// Mitsubishi GX Works2 project: KotelnyaPLC   PLC: FX3U/FX3UC (continued)
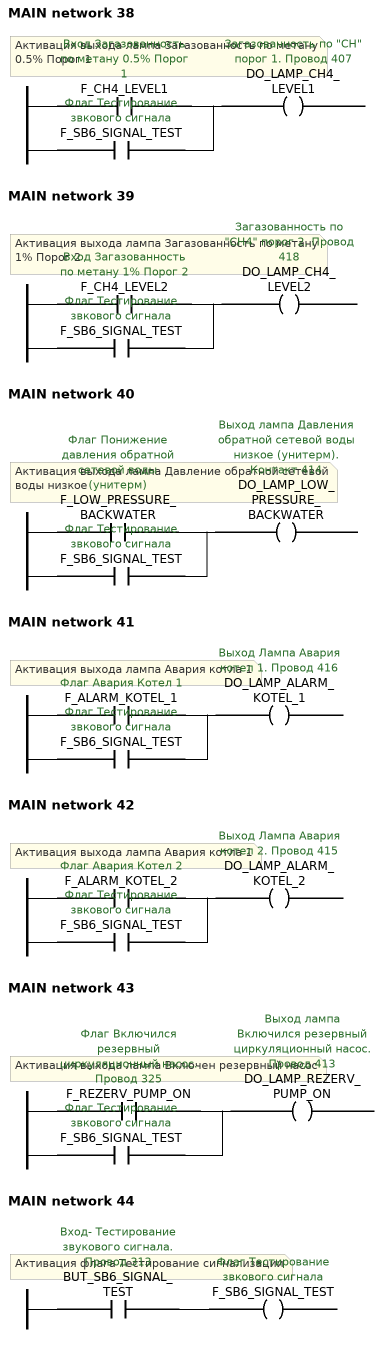
(* [picture p5: structured ladder/FBD of MAIN, networks 38 to 44] *)
(* network 38 *)
(* Активация выхода лампа Загазованность по метану 0.5% Порог 1 *)
DO_LAMP_CH4_LEVEL1 := F_CH4_LEVEL1 OR F_SB6_SIGNAL_TEST;
(* network 39 *)
(* Активация выхода лампа Загазованность по метану 1% Порог 2 *)
DO_LAMP_CH4_LEVEL2 := F_CH4_LEVEL2 OR F_SB6_SIGNAL_TEST;
(* network 40 *)
(* Активация выхода лампа Давление обратной сетевой воды низкое *)
DO_LAMP_LOW_PRESSURE_BACKWATER := F_LOW_PRESSURE_BACKWATER OR F_SB6_SIGNAL_TEST;
(* network 41 *)
(* Активация выхода лампа Авария котла 1 *)
DO_LAMP_ALARM_KOTEL_1 := F_ALARM_KOTEL_1 OR F_SB6_SIGNAL_TEST;
(* network 42 *)
(* Активация выхода лампа Авария котла 1 *)
DO_LAMP_ALARM_KOTEL_2 := F_ALARM_KOTEL_2 OR F_SB6_SIGNAL_TEST;
(* network 43 *)
(* Активация выхода лампа Включен резервный насос *)
DO_LAMP_REZERV_PUMP_ON := F_REZERV_PUMP_ON OR F_SB6_SIGNAL_TEST;
(* network 44 *)
(* Активация флага Тестирование сигнализации *)
F_SB6_SIGNAL_TEST := BUT_SB6_SIGNAL_TEST;
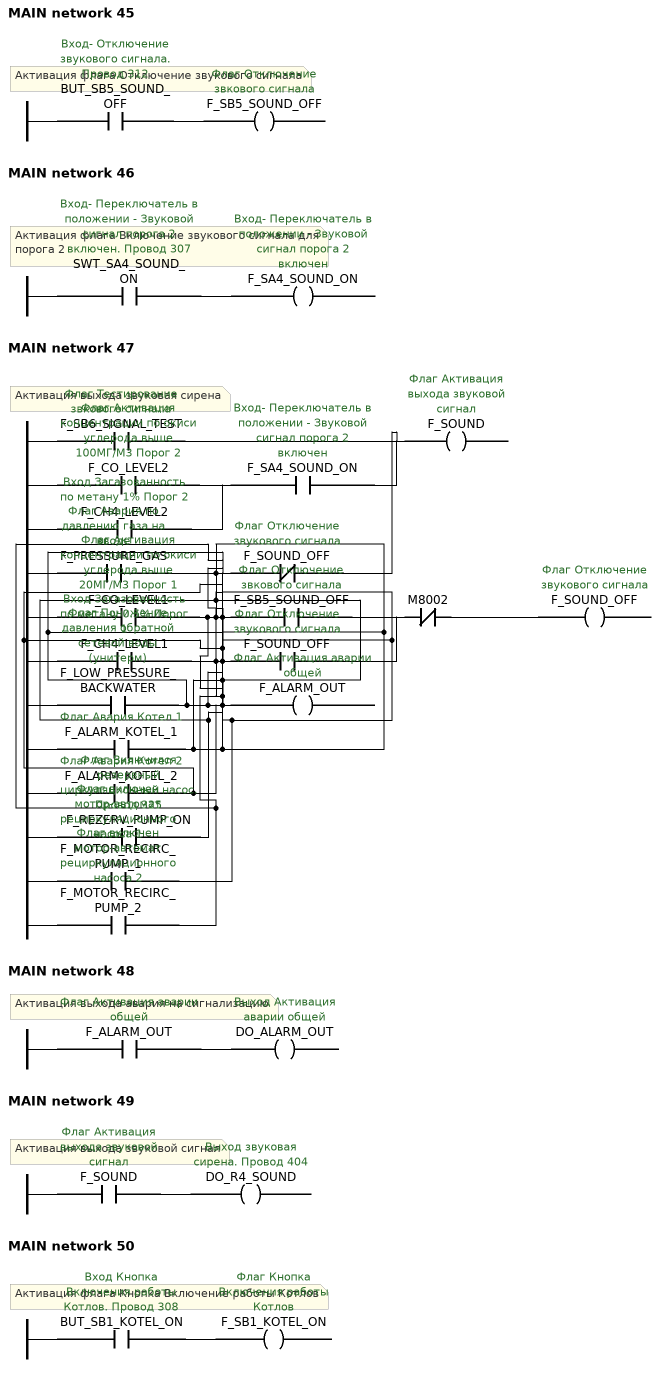
(* network 45 *)
(* Активация флага Отключение звукового сигнала *)
F_SB5_SOUND_OFF := BUT_SB5_SOUND_OFF;
(* network 46 *)
(* Активация флага Включение звукового сигнала для порога 2 *)
F_SA4_SOUND_ON := SWT_SA4_SOUND_ON;
(* network 47 *)
(* Активация выхода звуковая сирена *)
_p1 := F_PRESSURE_GAS OR F_CO_LEVEL1 OR F_CH4_LEVEL1 OR F_LOW_PRESSURE_BACKWATER OR F_ALARM_KOTEL_1 OR F_ALARM_KOTEL_2 OR F_REZERV_PUMP_ON OR F_MOTOR_RECIRC_PUMP_1 OR F_MOTOR_RECIRC_PUMP_2;
F_SOUND := F_SB6_SIGNAL_TEST OR ((F_CO_LEVEL2 OR F_CH4_LEVEL2) AND F_SA4_SOUND_ON) OR (_p1 AND NOT F_SOUND_OFF);
F_SOUND_OFF := ((_p1 AND F_SB5_SOUND_OFF) OR (_p1 AND F_SOUND_OFF)) AND NOT M8002;
F_ALARM_OUT := _p1;
(* network 48 *)
(* Активация выхода авария на сигнализацию *)
DO_ALARM_OUT := F_ALARM_OUT;
(* network 49 *)
(* Активация выхода звуковой сигнал *)
DO_R4_SOUND := F_SOUND;
(* network 50 *)
(* Активация флага Кнопка Включение работы Котлов *)
F_SB1_KOTEL_ON := BUT_SB1_KOTEL_ON;
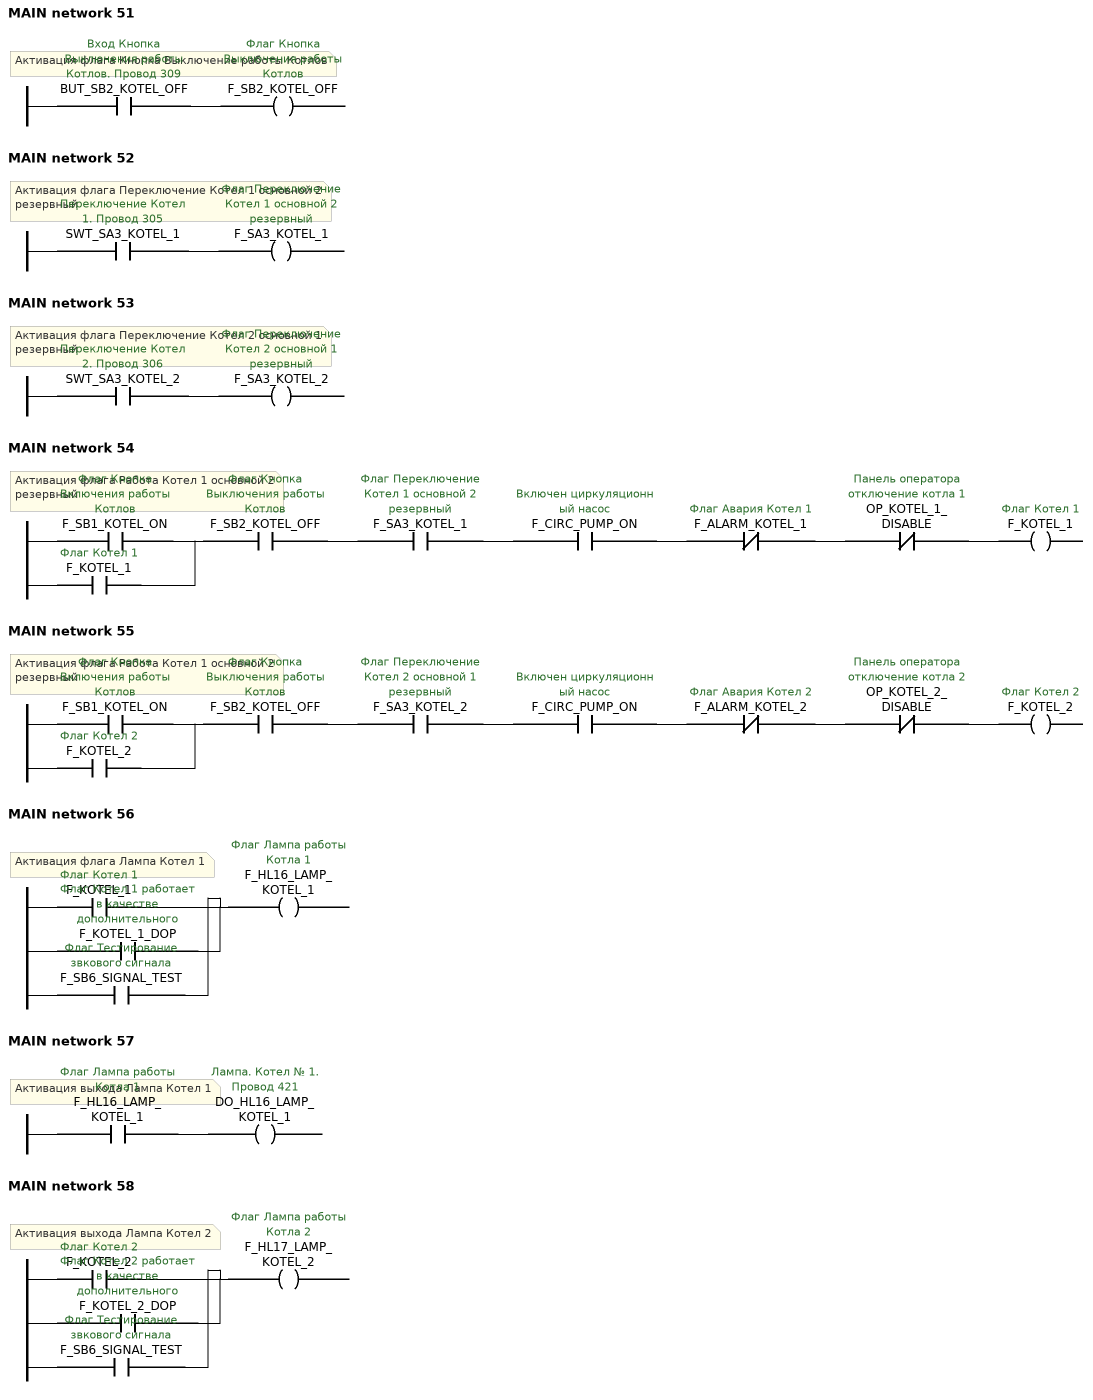
(* network 51 *)
(* Активация флага Кнопка Выключение работы Котлов *)
F_SB2_KOTEL_OFF := BUT_SB2_KOTEL_OFF;
(* network 52 *)
(* Активация флага Переключение Котел 1 основной 2 резервный *)
F_SA3_KOTEL_1 := SWT_SA3_KOTEL_1;
(* network 53 *)
(* Активация флага Переключение Котел 2 основной 1 резервный *)
F_SA3_KOTEL_2 := SWT_SA3_KOTEL_2;
(* network 54 *)
(* Активация флага Работа Котел 1 основной 2 резервный *)
F_KOTEL_1 := (((((F_SB1_KOTEL_ON OR F_KOTEL_1) AND F_SB2_KOTEL_OFF) AND F_SA3_KOTEL_1) AND F_CIRC_PUMP_ON) AND NOT F_ALARM_KOTEL_1) AND NOT OP_KOTEL_1_DISABLE;
(* network 55 *)
(* Активация флага Работа Котел 1 основной 2 резервный *)
F_KOTEL_2 := (((((F_SB1_KOTEL_ON OR F_KOTEL_2) AND F_SB2_KOTEL_OFF) AND F_SA3_KOTEL_2) AND F_CIRC_PUMP_ON) AND NOT F_ALARM_KOTEL_2) AND NOT OP_KOTEL_2_DISABLE;
(* network 56 *)
(* Активация флага Лампа Котел 1 *)
F_HL16_LAMP_KOTEL_1 := F_KOTEL_1 OR F_KOTEL_1_DOP OR F_SB6_SIGNAL_TEST;
(* network 57 *)
(* Активация выхода Лампа Котел 1 *)
DO_HL16_LAMP_KOTEL_1 := F_HL16_LAMP_KOTEL_1;
(* network 58 *)
(* Активация выхода Лампа Котел 2 *)
F_HL17_LAMP_KOTEL_2 := F_KOTEL_2 OR F_KOTEL_2_DOP OR F_SB6_SIGNAL_TEST;
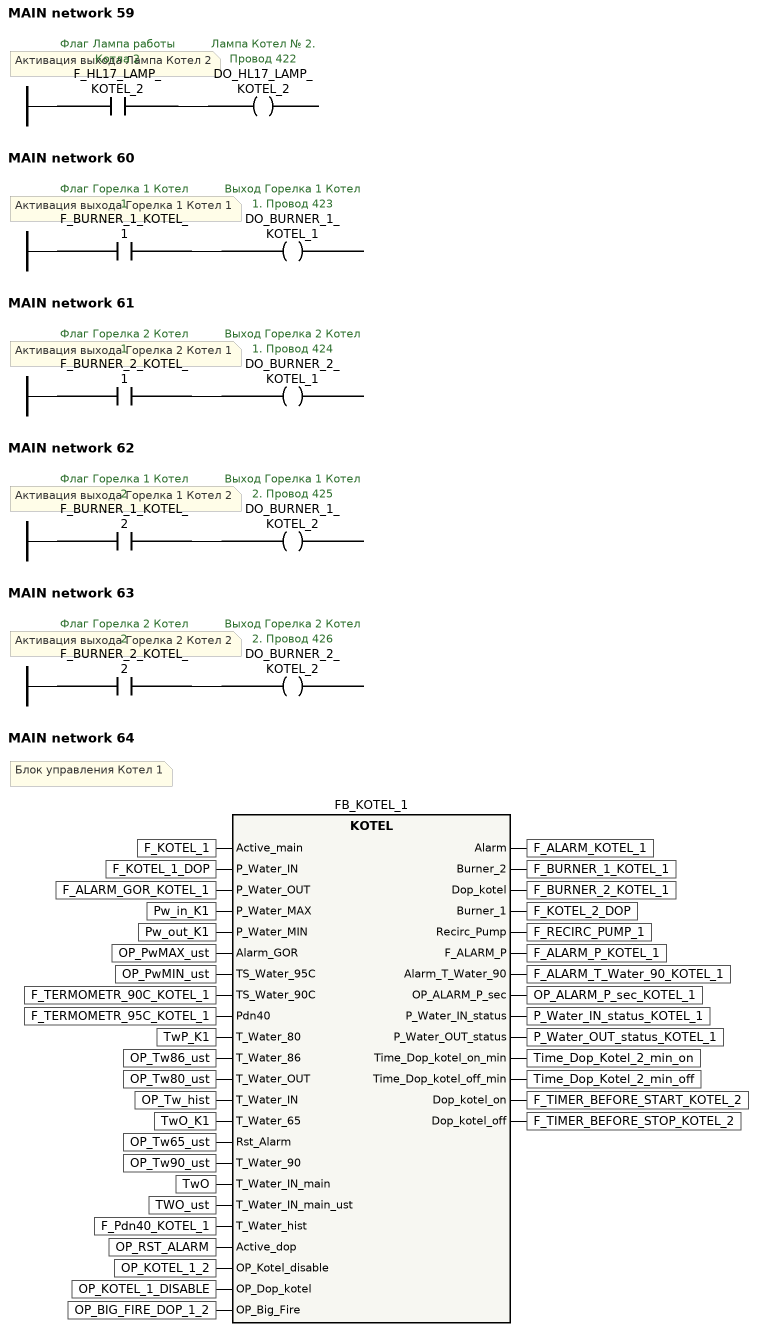
(* network 59 *)
(* Активация выхода Лампа Котел 2 *)
DO_HL17_LAMP_KOTEL_2 := F_HL17_LAMP_KOTEL_2;
(* network 60 *)
(* Активация выхода Горелка 1 Котел 1 *)
DO_BURNER_1_KOTEL_1 := F_BURNER_1_KOTEL_1;
(* network 61 *)
(* Активация выхода Горелка 2 Котел 1 *)
DO_BURNER_2_KOTEL_1 := F_BURNER_2_KOTEL_1;
(* network 62 *)
(* Активация выхода Горелка 1 Котел 2 *)
DO_BURNER_1_KOTEL_2 := F_BURNER_1_KOTEL_2;
(* network 63 *)
(* Активация выхода Горелка 2 Котел 2 *)
DO_BURNER_2_KOTEL_2 := F_BURNER_2_KOTEL_2;
(* network 64 *)
(* Блок управления Котел 1 *)
FB_KOTEL_1(Active_main := F_KOTEL_1, P_Water_IN := F_KOTEL_1_DOP, P_Water_OUT := F_ALARM_GOR_KOTEL_1, P_Water_MAX := Pw_in_K1, P_Water_MIN := Pw_out_K1, Alarm_GOR := OP_PwMAX_ust, TS_Water_95C := OP_PwMIN_ust, TS_Water_90C := F_TERMOMETR_90C_KOTEL_1, Pdn40 := F_TERMOMETR_95C_KOTEL_1, T_Water_80 := TwP_K1, T_Water_86 := OP_Tw86_ust, T_Water_OUT := OP_Tw80_ust, T_Water_IN := OP_Tw_hist, T_Water_65 := TwO_K1, Rst_Alarm := OP_Tw65_ust, T_Water_90 := OP_Tw90_ust, T_Water_IN_main := TwO, T_Water_IN_main_ust := TWO_ust, T_Water_hist := F_Pdn40_KOTEL_1, Active_dop := OP_RST_ALARM, OP_Kotel_disable := OP_KOTEL_1_2, OP_Dop_kotel := OP_KOTEL_1_DISABLE, OP_Big_Fire := OP_BIG_FIRE_DOP_1_2, Alarm => F_ALARM_KOTEL_1, Burner_2 => F_BURNER_1_KOTEL_1, Dop_kotel => F_BURNER_2_KOTEL_1, Burner_1 => F_KOTEL_2_DOP, Recirc_Pump => F_RECIRC_PUMP_1, F_ALARM_P => F_ALARM_P_KOTEL_1, Alarm_T_Water_90 => F_ALARM_T_Water_90_KOTEL_1, OP_ALARM_P_sec => OP_ALARM_P_sec_KOTEL_1, P_Water_IN_status => P_Water_IN_status_KOTEL_1, P_Water_OUT_status => P_Water_OUT_status_KOTEL_1, Time_Dop_kotel_on_min => Time_Dop_Kotel_2_min_on, Time_Dop_kotel_off_min => Time_Dop_Kotel_2_min_off, Dop_kotel_on => F_TIMER_BEFORE_START_KOTEL_2, Dop_kotel_off => F_TIMER_BEFORE_STOP_KOTEL_2);
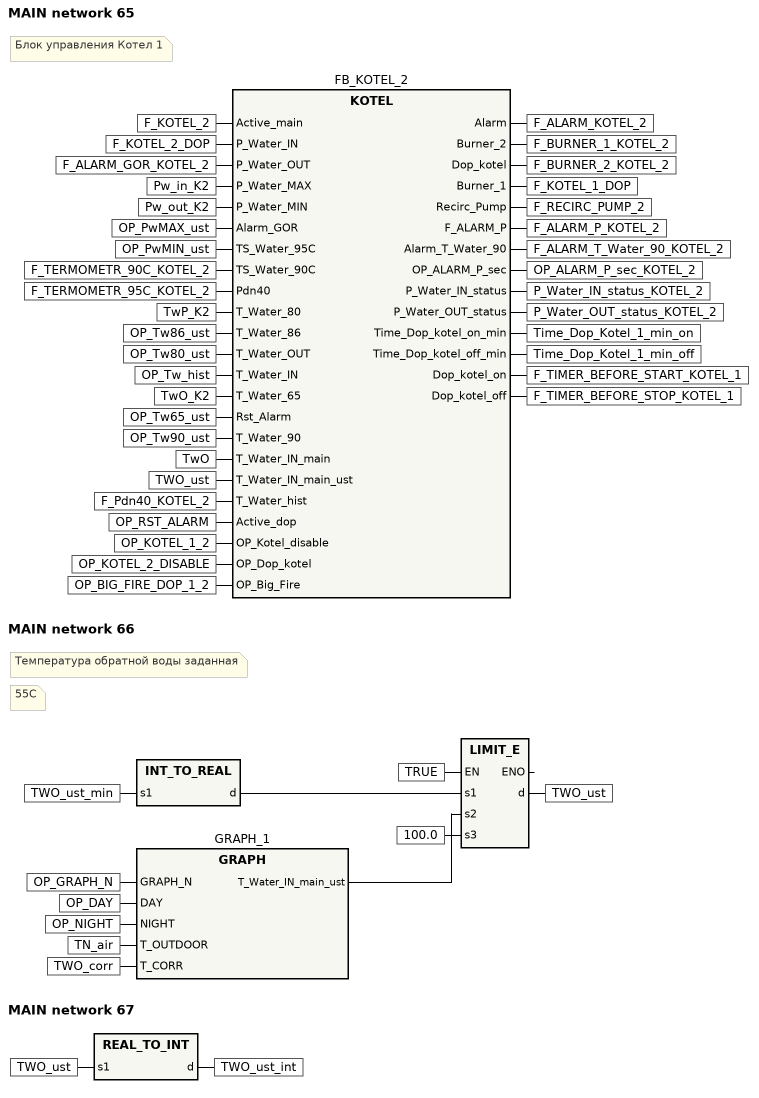
(* network 65 *)
(* Блок управления Котел 1 *)
FB_KOTEL_2(Active_main := F_KOTEL_2, P_Water_IN := F_KOTEL_2_DOP, P_Water_OUT := F_ALARM_GOR_KOTEL_2, P_Water_MAX := Pw_in_K2, P_Water_MIN := Pw_out_K2, Alarm_GOR := OP_PwMAX_ust, TS_Water_95C := OP_PwMIN_ust, TS_Water_90C := F_TERMOMETR_90C_KOTEL_2, Pdn40 := F_TERMOMETR_95C_KOTEL_2, T_Water_80 := TwP_K2, T_Water_86 := OP_Tw86_ust, T_Water_OUT := OP_Tw80_ust, T_Water_IN := OP_Tw_hist, T_Water_65 := TwO_K2, Rst_Alarm := OP_Tw65_ust, T_Water_90 := OP_Tw90_ust, T_Water_IN_main := TwO, T_Water_IN_main_ust := TWO_ust, T_Water_hist := F_Pdn40_KOTEL_2, Active_dop := OP_RST_ALARM, OP_Kotel_disable := OP_KOTEL_1_2, OP_Dop_kotel := OP_KOTEL_2_DISABLE, OP_Big_Fire := OP_BIG_FIRE_DOP_1_2, Alarm => F_ALARM_KOTEL_2, Burner_2 => F_BURNER_1_KOTEL_2, Dop_kotel => F_BURNER_2_KOTEL_2, Burner_1 => F_KOTEL_1_DOP, Recirc_Pump => F_RECIRC_PUMP_2, F_ALARM_P => F_ALARM_P_KOTEL_2, Alarm_T_Water_90 => F_ALARM_T_Water_90_KOTEL_2, OP_ALARM_P_sec => OP_ALARM_P_sec_KOTEL_2, P_Water_IN_status => P_Water_IN_status_KOTEL_2, P_Water_OUT_status => P_Water_OUT_status_KOTEL_2, Time_Dop_kotel_on_min => Time_Dop_Kotel_1_min_on, Time_Dop_kotel_off_min => Time_Dop_Kotel_1_min_off, Dop_kotel_on => F_TIMER_BEFORE_START_KOTEL_1, Dop_kotel_off => F_TIMER_BEFORE_STOP_KOTEL_1);
(* network 66 *)
(* Температура обратной воды заданная *)
(* 55C *)
GRAPH_1(GRAPH_N := OP_GRAPH_N, DAY := OP_DAY, NIGHT := OP_NIGHT, T_OUTDOOR := TN_air, T_CORR := TWO_corr);
LIMIT_E(TRUE, INT_TO_REAL(TWO_ust_min), GRAPH_1.T_Water_IN_main_ust, 100.0, TWO_ust);
(* network 67 *)
TWO_ust_int := REAL_TO_INT(TWO_ust);
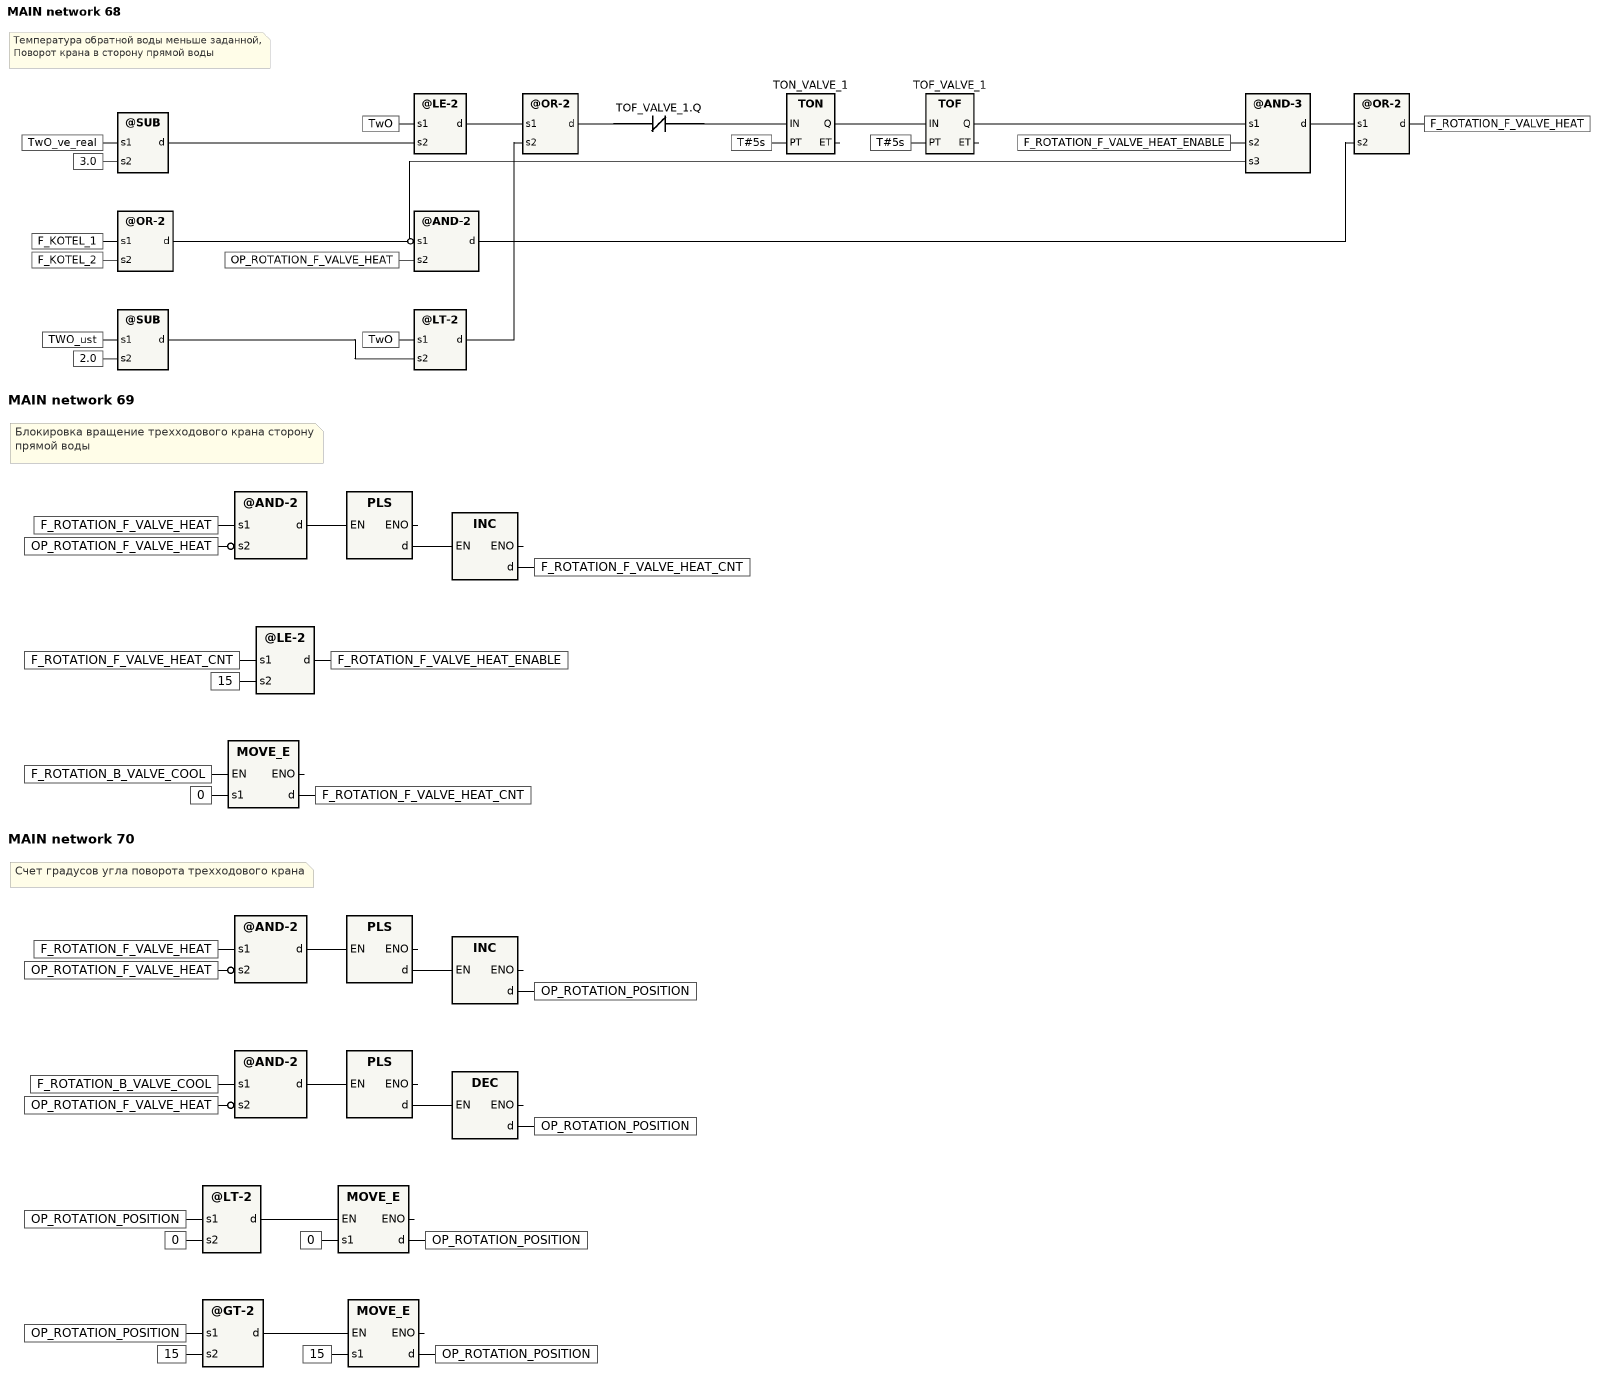
(* network 68 *)
(* Температура обратной воды меньше заданной, Поворот крана в сторону прямой воды *)
TON_VALVE_1(IN := @OR-2(@LE-2(TwO, @SUB(TwO_ve_real, 3.0)), @LT-2(TwO, @SUB(TWO_ust, 2.0))) AND NOT TOF_VALVE_1.Q, PT := T#5s);
TOF_VALVE_1(IN := TON_VALVE_1.Q, PT := T#5s);
_p1 := @OR-2(F_KOTEL_1, F_KOTEL_2);
F_ROTATION_F_VALVE_HEAT := @OR-2(@AND-3(TOF_VALVE_1.Q, F_ROTATION_F_VALVE_HEAT_ENABLE, _p1), @AND-2(NOT _p1, OP_ROTATION_F_VALVE_HEAT));
(* network 69 *)
(* Блокировка вращение трехходового крана сторону прямой воды *)
PLS(@AND-2(F_ROTATION_F_VALVE_HEAT, NOT OP_ROTATION_F_VALVE_HEAT), _t1);
INC(_t1, F_ROTATION_F_VALVE_HEAT_CNT);
F_ROTATION_F_VALVE_HEAT_ENABLE := @LE-2(F_ROTATION_F_VALVE_HEAT_CNT, 15);
MOVE_E(F_ROTATION_B_VALVE_COOL, 0, F_ROTATION_F_VALVE_HEAT_CNT);
(* network 70 *)
(* Счет градусов угла поворота трехходового крана *)
PLS(@AND-2(F_ROTATION_F_VALVE_HEAT, NOT OP_ROTATION_F_VALVE_HEAT), _t1);
INC(_t1, OP_ROTATION_POSITION);
PLS(@AND-2(F_ROTATION_B_VALVE_COOL, NOT OP_ROTATION_F_VALVE_HEAT), _t2);
DEC(_t2, OP_ROTATION_POSITION);
MOVE_E(@LT-2(OP_ROTATION_POSITION, 0), 0, OP_ROTATION_POSITION);
MOVE_E(@GT-2(OP_ROTATION_POSITION, 15), 15, OP_ROTATION_POSITION);
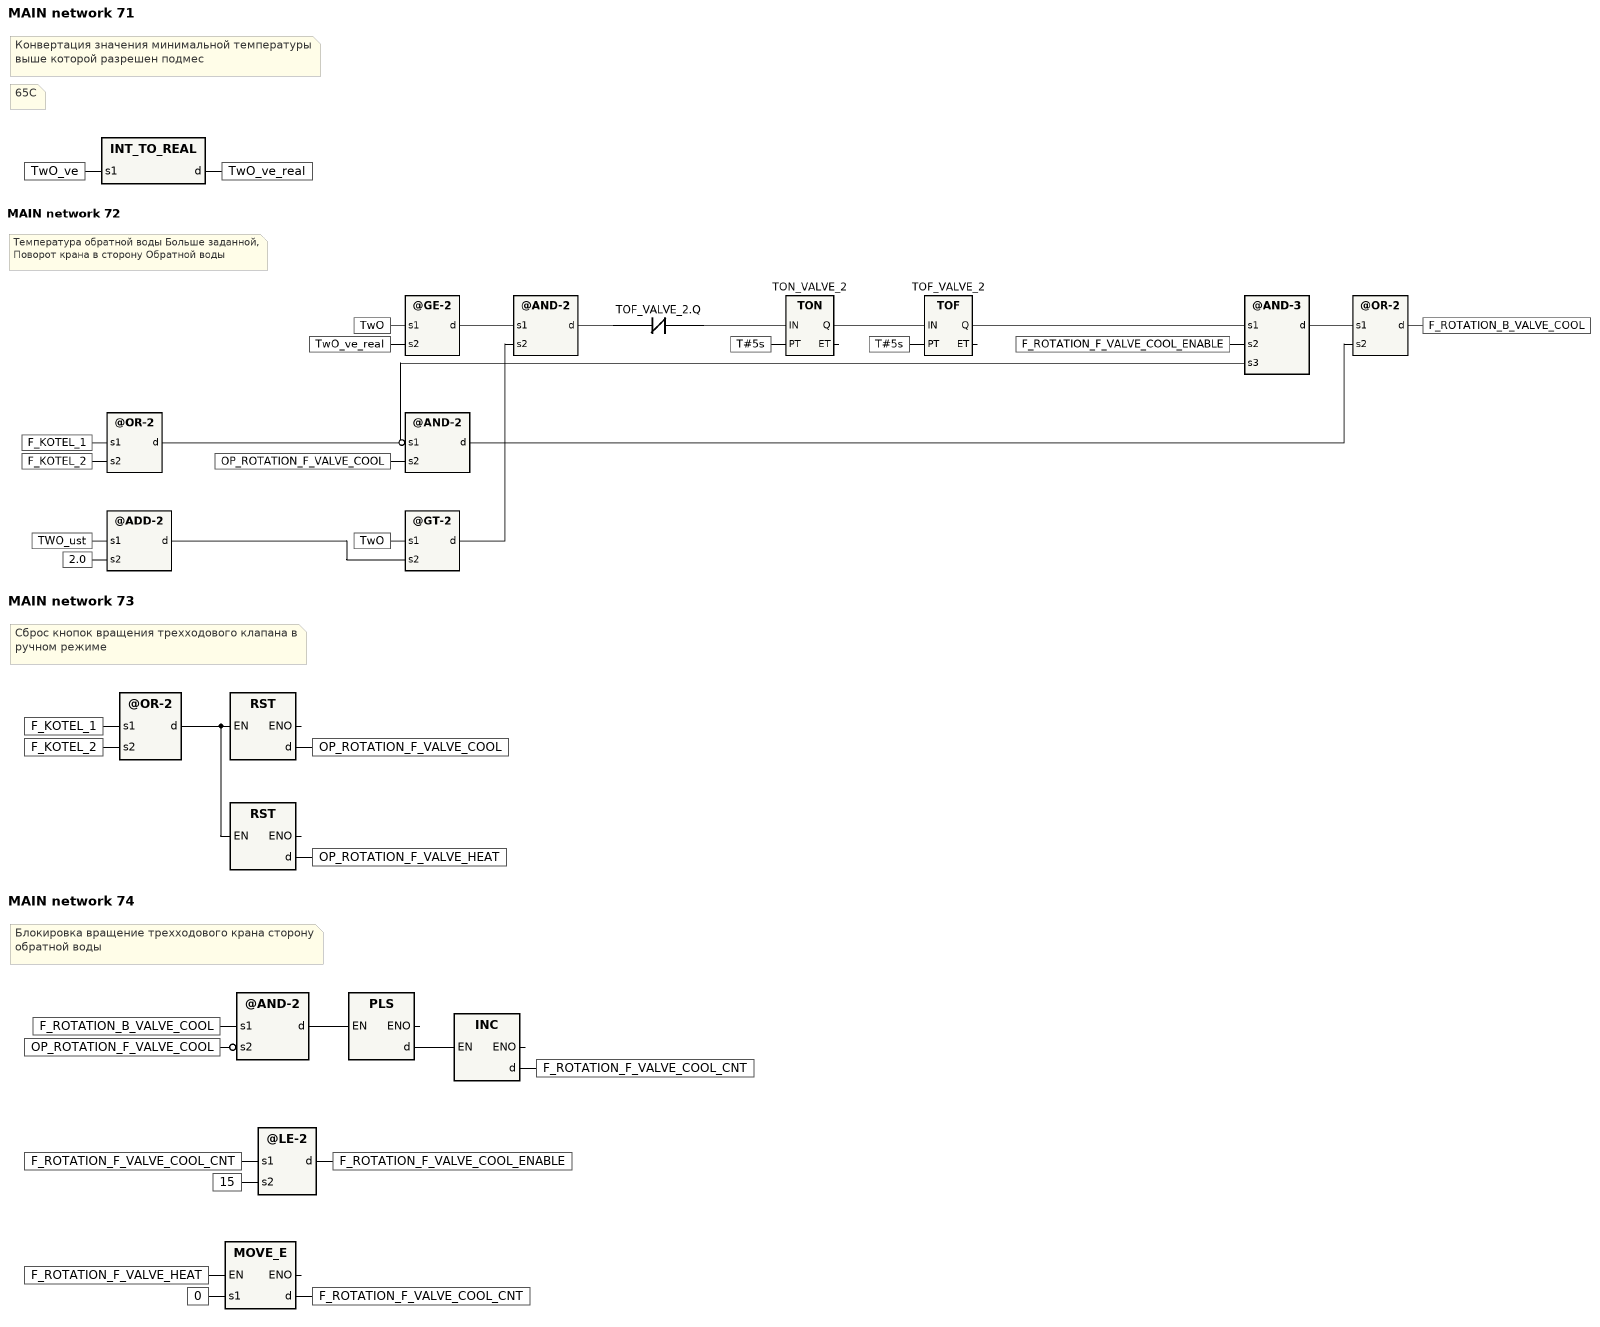
(* network 71 *)
(* Конвертация значения минимальной температуры выше которой разрешен подмес *)
(* 65С *)
TwO_ve_real := INT_TO_REAL(TwO_ve);
(* network 72 *)
(* Температура обратной воды Больше заданной, Поворот крана в сторону Обратной воды *)
TON_VALVE_2(IN := @AND-2(@GE-2(TwO, TwO_ve_real), @GT-2(TwO, @ADD-2(TWO_ust, 2.0))) AND NOT TOF_VALVE_2.Q, PT := T#5s);
TOF_VALVE_2(IN := TON_VALVE_2.Q, PT := T#5s);
_p1 := @OR-2(F_KOTEL_1, F_KOTEL_2);
F_ROTATION_B_VALVE_COOL := @OR-2(@AND-3(TOF_VALVE_2.Q, F_ROTATION_F_VALVE_COOL_ENABLE, _p1), @AND-2(NOT _p1, OP_ROTATION_F_VALVE_COOL));
(* network 73 *)
(* Сброс кнопок вращения трехходового клапана в ручном режиме *)
_p1 := @OR-2(F_KOTEL_1, F_KOTEL_2);
RST(_p1, OP_ROTATION_F_VALVE_COOL);
RST(_p1, OP_ROTATION_F_VALVE_HEAT);
(* network 74 *)
(* Блокировка вращение трехходового крана сторону обратной воды *)
PLS(@AND-2(F_ROTATION_B_VALVE_COOL, NOT OP_ROTATION_F_VALVE_COOL), _t1);
INC(_t1, F_ROTATION_F_VALVE_COOL_CNT);
F_ROTATION_F_VALVE_COOL_ENABLE := @LE-2(F_ROTATION_F_VALVE_COOL_CNT, 15);
MOVE_E(F_ROTATION_F_VALVE_HEAT, 0, F_ROTATION_F_VALVE_COOL_CNT);
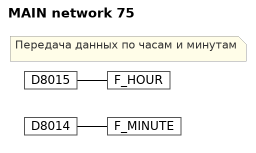
(* network 75 *)
(* Передача данных по часам и минутам *)
F_HOUR := D8015;
F_MINUTE := D8014;
END_PROGRAM

PROGRAM AIN_FBD
VAR
  FX2N_8AD_1 : FX2N_8AD;
  Reset_8AD : BOOL;
  AnalogInputCh1_8AD : INT;  (* Провод 355 *)
  AnalogInputCh2_8AD : INT;  (* Провод 356 *)
  AnalogInputCh3_8AD : INT;  (* Провод 357 *)
  AnalogInputCh4_8AD : INT;  (* Провод 358 *)
  AnalogInputCh5_8AD : INT;  (* Провод 359 *)
  AnalogInputCh6_8AD : INT;  (* Провод 360 *)
  AnalogInputCh7_8AD : INT;  (* Провод 361 *)
  AnalogInputCh8_8AD : INT;  (* Провод 362 *)
  GeneralError_8AD : BOOL;
  RangeError_8AD : BOOL;
  ErrorStatusDetails_8AD : WORD;
  ScaleOverStatus_8AD : WORD;
  ConversionActive_8AD : BOOL;
  FX2N_4AD_1 : FX2N_4AD;
  ConversionActive_4AD_1 : BOOL;
  AnalogInputPresentCh1_4AD_1 : INT;  (* Провод 363 *)
  AnalogInputPresentCh2_4AD_1 : INT;  (* Провод 364 *)
  AnalogInputPresentCh3_4AD_1 : INT;  (* Провод 365 *)
  AnalogInputPresentCh4_4AD_1 : INT;  (* Провод 366 *)
  AnalogInputAvgCh1_4AD_1 : INT;
  AnalogInputAvgCh2_4AD_1 : INT;
  AnalogInputAvgCh3_4AD_1 : INT;
  AnalogInputAvgCh4_4AD_1 : INT;
  GeneralError_4AD_1 : BOOL;
  RangeError_4AD_1 : BOOL;
  AverageError_4AD_1 : BOOL;
  Sensor_1_converter : 4-20mA_TO_VALUE;
  Sensor_2_converter : 4-20mA_TO_VALUE;
  Sensor_4_converter : 4-20mA_TO_VALUE;
  Sensor_3_converter : 4-20mA_TO_VALUE;
  Sensor_5_converter : 4-20mA_TO_VALUE;
  Sensor_6_converter : 4-20mA_TO_VALUE;
  Sensor_7_converter : 4-20mA_TO_VALUE;
  Sensor_8_converter : 4-20mA_TO_VALUE;
  Sensor_9_converter : 4-20mA_TO_VALUE;
  Sensor_10_converter : 4-20mA_TO_VALUE;
  Sensor_11_converter : 4-20mA_TO_VALUE;
  Sensor_12_converter : 4-20mA_TO_VALUE;
  FX2N_4AD_2 : FX2N_4AD;
  ConversionActive_4AD_2 : BOOL;
  AnalogInputPresentCh1_4AD_2 : INT;  (* Провод 363 *)
  AnalogInputPresentCh2_4AD_2 : INT;  (* Провод 364 *)
  AnalogInputPresentCh3_4AD_2 : INT;  (* Провод 365 *)
  AnalogInputPresentCh4_4AD_2 : INT;  (* Провод 366 *)
  AnalogInputAvgCh1_4AD_2 : INT;
  AnalogInputAvgCh2_4AD_2 : INT;
  AnalogInputAvgCh3_4AD_2 : INT;
  AnalogInputAvgCh4_4AD_2 : INT;
  GeneralError_4AD_2 : BOOL;
  RangeError_4AD_2 : BOOL;
  AverageError_4AD_2 : BOOL;
  Sensor_13_converter : 4-20mA_TO_VALUE;
  Sensor_14_converter : 4-20mA_TO_VALUE;
END_VAR
(* structured ladder/FBD written out as ST: instructions are called as NAME(EN, inputs, outputs); _pN, _eN, _tN stand for wires *)
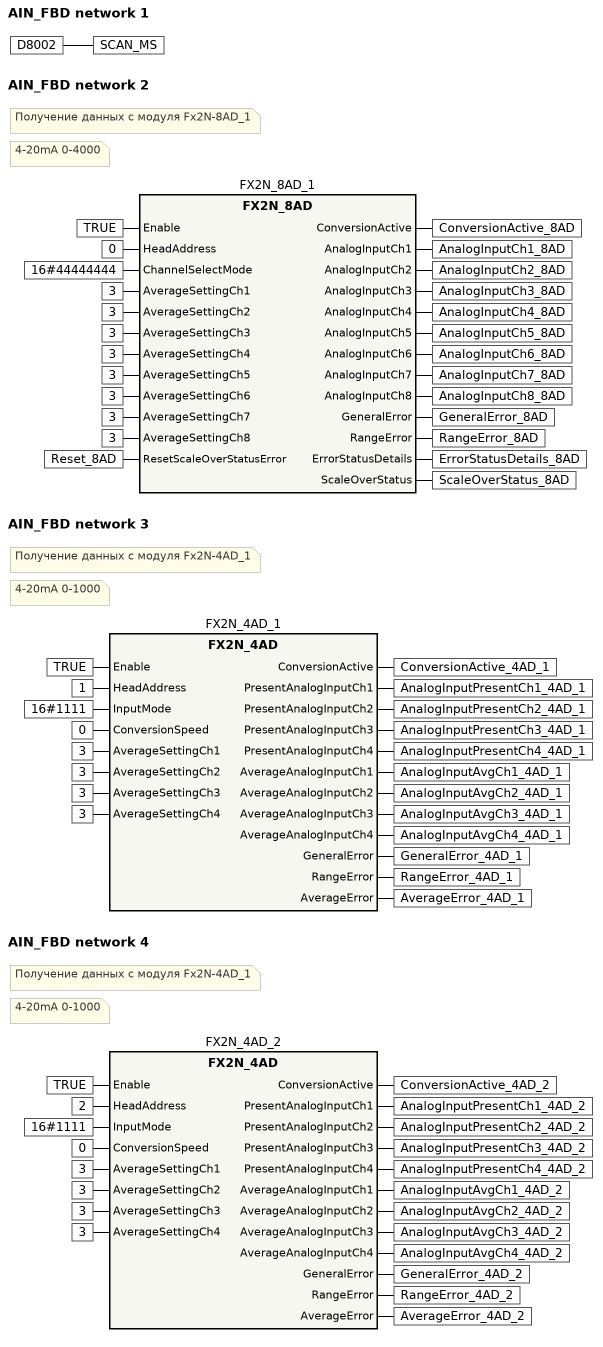
(* network 1 *)
SCAN_MS := D8002;
(* network 2 *)
(* Получение данных с модуля Fx2N-8AD_1 *)
(* 4-20mA 0-4000 *)
FX2N_8AD_1(Enable := TRUE, HeadAddress := 0, ChannelSelectMode := 16#44444444, AverageSettingCh1 := 3, AverageSettingCh2 := 3, AverageSettingCh3 := 3, AverageSettingCh4 := 3, AverageSettingCh5 := 3, AverageSettingCh6 := 3, AverageSettingCh7 := 3, AverageSettingCh8 := 3, ResetScaleOverStatusError := Reset_8AD, ConversionActive => ConversionActive_8AD, AnalogInputCh1 => AnalogInputCh1_8AD, AnalogInputCh2 => AnalogInputCh2_8AD, AnalogInputCh3 => AnalogInputCh3_8AD, AnalogInputCh4 => AnalogInputCh4_8AD, AnalogInputCh5 => AnalogInputCh5_8AD, AnalogInputCh6 => AnalogInputCh6_8AD, AnalogInputCh7 => AnalogInputCh7_8AD, AnalogInputCh8 => AnalogInputCh8_8AD, GeneralError => GeneralError_8AD, RangeError => RangeError_8AD, ErrorStatusDetails => ErrorStatusDetails_8AD, ScaleOverStatus => ScaleOverStatus_8AD);
(* network 3 *)
(* Получение данных с модуля Fx2N-4AD_1 *)
(* 4-20mA 0-1000 *)
FX2N_4AD_1(Enable := TRUE, HeadAddress := 1, InputMode := 16#1111, ConversionSpeed := 0, AverageSettingCh1 := 3, AverageSettingCh2 := 3, AverageSettingCh3 := 3, AverageSettingCh4 := 3, ConversionActive => ConversionActive_4AD_1, PresentAnalogInputCh1 => AnalogInputPresentCh1_4AD_1, PresentAnalogInputCh2 => AnalogInputPresentCh2_4AD_1, PresentAnalogInputCh3 => AnalogInputPresentCh3_4AD_1, PresentAnalogInputCh4 => AnalogInputPresentCh4_4AD_1, AverageAnalogInputCh1 => AnalogInputAvgCh1_4AD_1, AverageAnalogInputCh2 => AnalogInputAvgCh2_4AD_1, AverageAnalogInputCh3 => AnalogInputAvgCh3_4AD_1, AverageAnalogInputCh4 => AnalogInputAvgCh4_4AD_1, GeneralError => GeneralError_4AD_1, RangeError => RangeError_4AD_1, AverageError => AverageError_4AD_1);
(* network 4 *)
(* Получение данных с модуля Fx2N-4AD_1 *)
(* 4-20mA 0-1000 *)
FX2N_4AD_2(Enable := TRUE, HeadAddress := 2, InputMode := 16#1111, ConversionSpeed := 0, AverageSettingCh1 := 3, AverageSettingCh2 := 3, AverageSettingCh3 := 3, AverageSettingCh4 := 3, ConversionActive => ConversionActive_4AD_2, PresentAnalogInputCh1 => AnalogInputPresentCh1_4AD_2, PresentAnalogInputCh2 => AnalogInputPresentCh2_4AD_2, PresentAnalogInputCh3 => AnalogInputPresentCh3_4AD_2, PresentAnalogInputCh4 => AnalogInputPresentCh4_4AD_2, AverageAnalogInputCh1 => AnalogInputAvgCh1_4AD_2, AverageAnalogInputCh2 => AnalogInputAvgCh2_4AD_2, AverageAnalogInputCh3 => AnalogInputAvgCh3_4AD_2, AverageAnalogInputCh4 => AnalogInputAvgCh4_4AD_2, GeneralError => GeneralError_4AD_2, RangeError => RangeError_4AD_2, AverageError => AverageError_4AD_2);